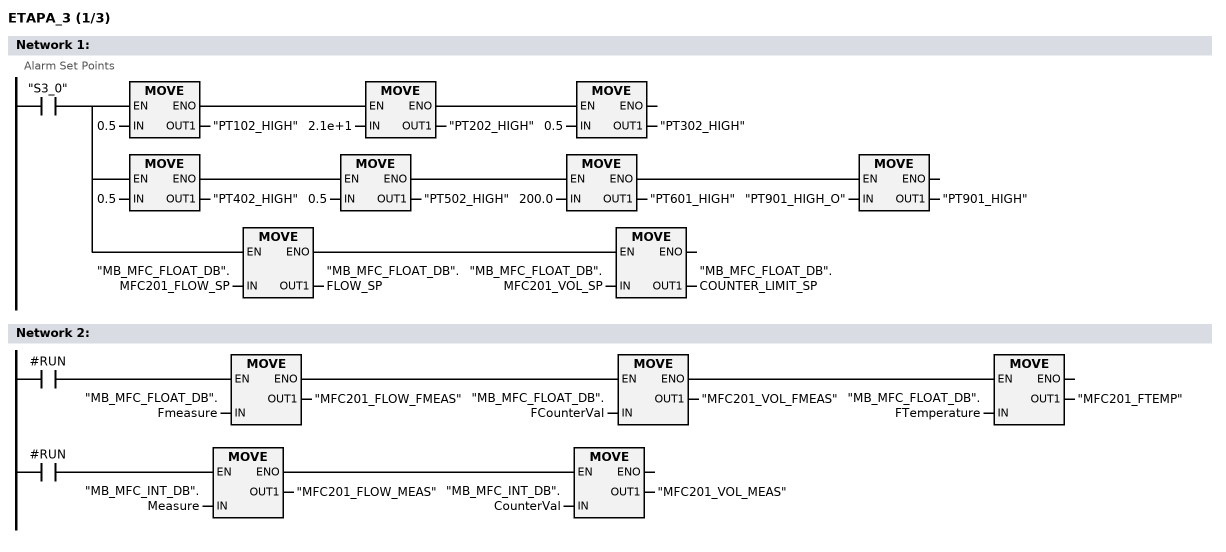
   RUNG wire#powerrail
      Contact( "S3_0" )
      wire#w1
      { S7_GenerateENO := "TRUE" } Move(in := 0.5, out1 => "PT102_HIGH")
      { S7_GenerateENO := "TRUE" } Move(in := 2.1e+1, out1 => "PT202_HIGH")
      { S7_GenerateENO := "TRUE" } Move(in := 0.5, out1 => "PT302_HIGH")
   END_RUNG
   RUNG wire#w1
      { S7_GenerateENO := "TRUE" } Move(in := 0.5, out1 => "PT402_HIGH")
      { S7_GenerateENO := "TRUE" } Move(in := 0.5, out1 => "PT502_HIGH")
      { S7_GenerateENO := "TRUE" } Move(in := 200.0, out1 => "PT601_HIGH")
      { S7_GenerateENO := "TRUE" } Move(in := "PT901_HIGH_O", out1 => "PT901_HIGH")
   END_RUNG
   RUNG wire#w1
      Move(in := "MB_MFC_FLOAT_DB".MFC201_FLOW_SP, out1 => "MB_MFC_FLOAT_DB".FLOW_SP)
      Move(in := "MB_MFC_FLOAT_DB".MFC201_VOL_SP, out1 => "MB_MFC_FLOAT_DB".COUNTER_LIMIT_SP)
   END_RUNG
   // the same network as SCL:
   // ENO of a box is taken as its EN; it also drops when the box reports an error
   IF "S3_0" THEN
       "PT102_HIGH" := 0.5;
       "PT202_HIGH" := 2.1e+1;
       "PT302_HIGH" := 0.5;
       "PT402_HIGH" := 0.5;
       "PT502_HIGH" := 0.5;
       "PT601_HIGH" := 200.0;
       "PT901_HIGH" := "PT901_HIGH_O";
       "MB_MFC_FLOAT_DB".FLOW_SP := "MB_MFC_FLOAT_DB".MFC201_FLOW_SP;
       "MB_MFC_FLOAT_DB".COUNTER_LIMIT_SP := "MB_MFC_FLOAT_DB".MFC201_VOL_SP;
   END_IF;
END_REGION

REGION Network 2
   RUNG wire#powerrail
      Contact( #RUN )
      { S7_GenerateENO := "TRUE" } Move(in := "MB_MFC_FLOAT_DB".Fmeasure, out1 => "MFC201_FLOW_FMEAS")
      { S7_GenerateENO := "TRUE" } Move(in := "MB_MFC_FLOAT_DB".FCounterVal, out1 => "MFC201_VOL_FMEAS")
      { S7_GenerateENO := "TRUE" } Move(in := "MB_MFC_FLOAT_DB".FTemperature, out1 => "MFC201_FTEMP")
   END_RUNG
   RUNG wire#powerrail
      Contact( #RUN )
      { S7_GenerateENO := "TRUE" } Move(in := "MB_MFC_INT_DB".Measure, out1 => "MFC201_FLOW_MEAS")
      { S7_GenerateENO := "TRUE" } Move(in := "MB_MFC_INT_DB".CounterVal, out1 => "MFC201_VOL_MEAS")
   END_RUNG
   // the same network as SCL:
   // ENO of a box is taken as its EN; it also drops when the box reports an error
   IF #RUN THEN
       "MFC201_FLOW_FMEAS" := "MB_MFC_FLOAT_DB".Fmeasure;
       "MFC201_VOL_FMEAS" := "MB_MFC_FLOAT_DB".FCounterVal;
       "MFC201_FTEMP" := "MB_MFC_FLOAT_DB".FTemperature;
       "MFC201_FLOW_MEAS" := "MB_MFC_INT_DB".Measure;
       "MFC201_VOL_MEAS" := "MB_MFC_INT_DB".CounterVal;
   END_IF;
END_REGION

REGION Network 3
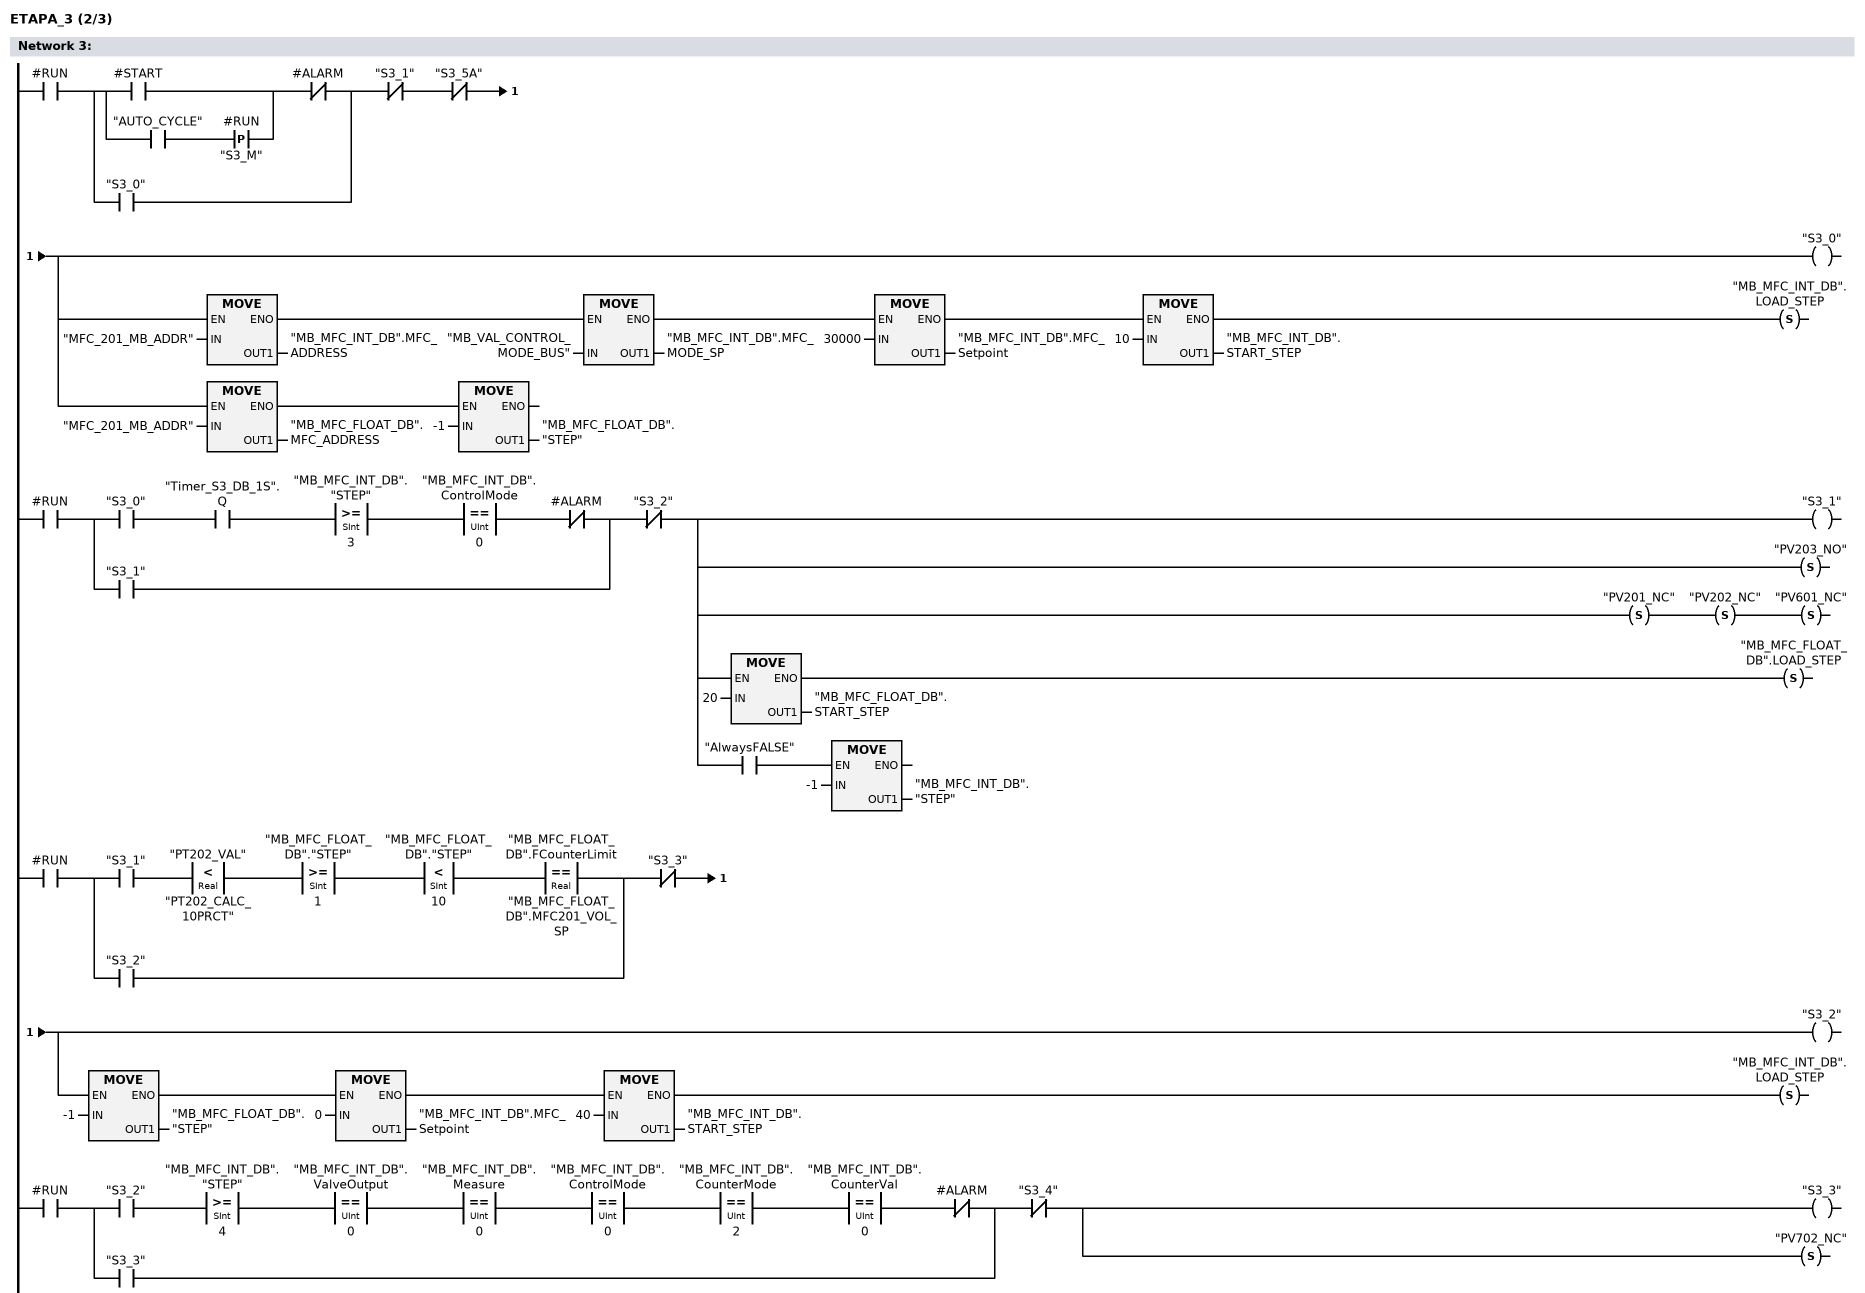
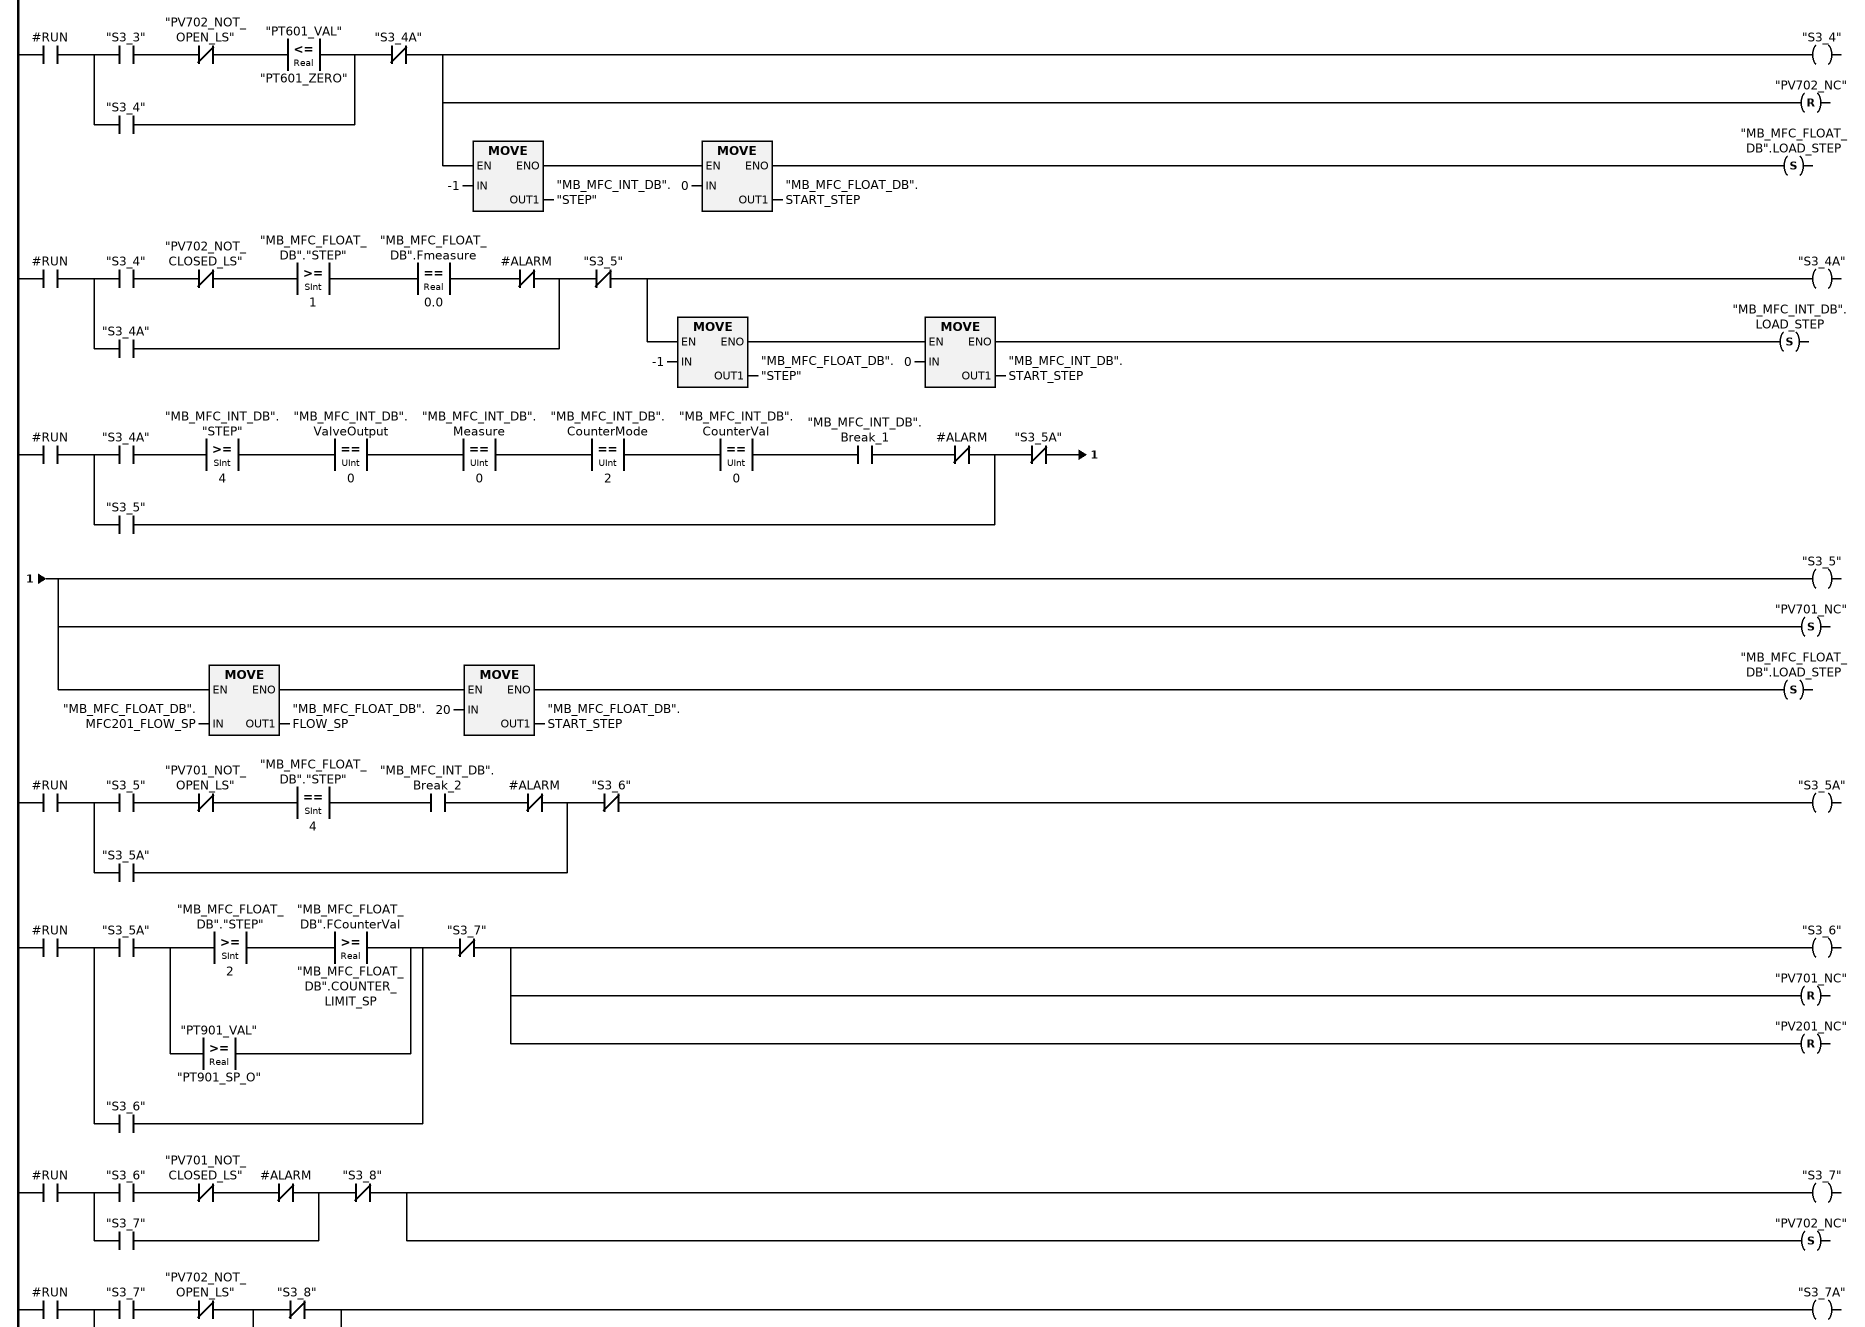
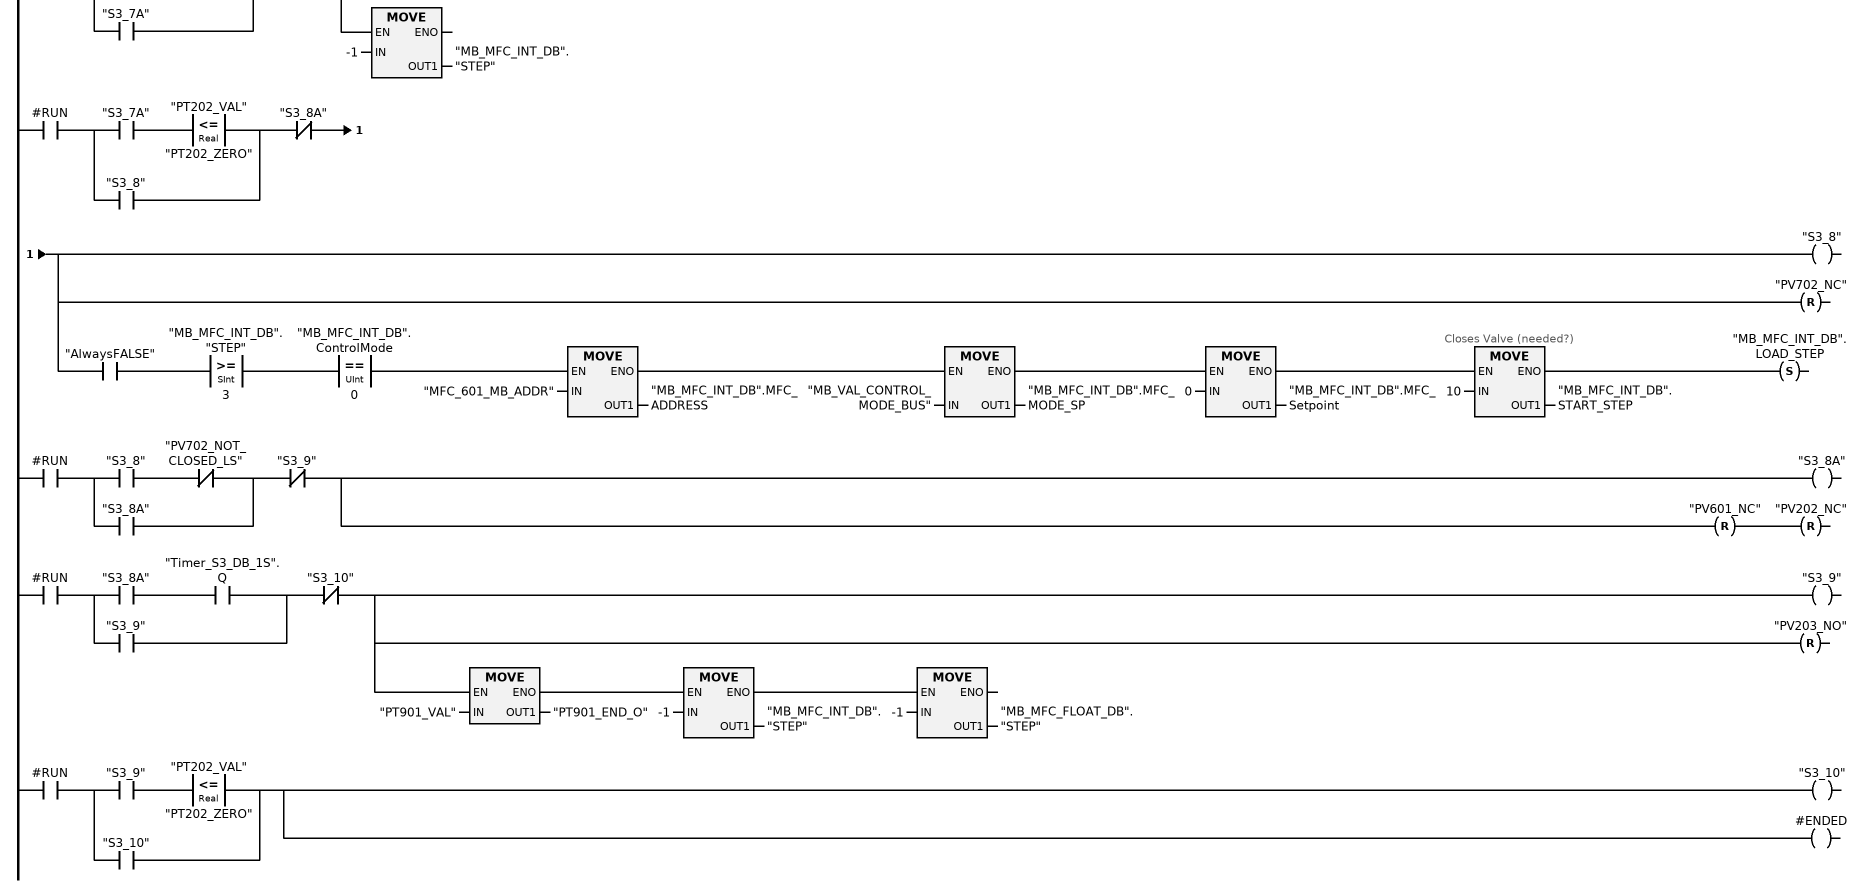
   RUNG wire#powerrail
      Contact( #RUN )
      wire#w1
      Contact( #START )
      wire#w2
      I_Contact( #ALARM )
      wire#w3
      I_Contact( "S3_1" )
      I_Contact( "S3_5A" )
      wire#w4
      Coil( "S3_0" )
   END_RUNG
   RUNG wire#w1
      Contact( "AUTO_CYCLE" )
      P_Contact(operand := #RUN, bit := "S3_M")
   END_RUNG wire#w2
   RUNG wire#w1
      Contact( "S3_0" )
   END_RUNG wire#w3
   RUNG wire#w4
      Move(in := "MFC_201_MB_ADDR", out1 => "MB_MFC_INT_DB".MFC_ADDRESS)
      Move(in := "MB_VAL_CONTROL_MODE_BUS", out1 => "MB_MFC_INT_DB".MFC_MODE_SP)
      Move(in := 30000, out1 => "MB_MFC_INT_DB".MFC_Setpoint)
      Move(in := 10, out1 => "MB_MFC_INT_DB".START_STEP)
      S_Coil( "MB_MFC_INT_DB".LOAD_STEP )
   END_RUNG
   RUNG wire#w4
      Move(in := "MFC_201_MB_ADDR", out1 => "MB_MFC_FLOAT_DB".MFC_ADDRESS)
      Move(in := -1, out1 => "MB_MFC_FLOAT_DB"."STEP")
   END_RUNG
   RUNG wire#powerrail
      Contact( #RUN )
      wire#w5
      Contact( "S3_0" )
      Contact( "Timer_S3_DB_1S".Q )
      { S7_Templates := "SrcType := SInt" } GE_Contact(in1 := "MB_MFC_INT_DB"."STEP", in2 := 3)
      { S7_Templates := "SrcType := UInt" } EQ_Contact(in1 := "MB_MFC_INT_DB".ControlMode, in2 := 0)
      I_Contact( #ALARM )
      wire#w6
      I_Contact( "S3_2" )
      wire#w7
      Coil( "S3_1" )
   END_RUNG
   RUNG wire#w5
      Contact( "S3_1" )
   END_RUNG wire#w6
   RUNG wire#w7
      S_Coil( "PV203_NO" )
   END_RUNG
   RUNG wire#w7
      S_Coil( "PV201_NC" )
      S_Coil( "PV202_NC" )
      S_Coil( "PV601_NC" )
   END_RUNG
   RUNG wire#w7
      Move(in := 20, out1 => "MB_MFC_FLOAT_DB".START_STEP)
      S_Coil( "MB_MFC_FLOAT_DB".LOAD_STEP )
   END_RUNG
   RUNG wire#w7
      Contact( "AlwaysFALSE" )
      Move(in := -1, out1 => "MB_MFC_INT_DB"."STEP")
   END_RUNG
   RUNG wire#powerrail
      Contact( #RUN )
      wire#w8
      Contact( "S3_1" )
      { S7_Templates := "SrcType := Real" } LT_Contact(in1 := "PT202_VAL", in2 := "PT202_CALC_10PRCT")
      { S7_Templates := "SrcType := SInt" } GE_Contact(in1 := "MB_MFC_FLOAT_DB"."STEP", in2 := 1)
      { S7_Templates := "SrcType := SInt" } LT_Contact(in1 := "MB_MFC_FLOAT_DB"."STEP", in2 := 10)
      { S7_Templates := "SrcType := Real" } EQ_Contact(in1 := "MB_MFC_FLOAT_DB".FCounterLimit, in2 := "MB_MFC_FLOAT_DB".MFC201_VOL_SP)
      wire#w9
      I_Contact( "S3_3" )
      wire#w10
      Coil( "S3_2" )
   END_RUNG
   RUNG wire#w8
      Contact( "S3_2" )
   END_RUNG wire#w9
   RUNG wire#w10
      Move(in := -1, out1 => "MB_MFC_FLOAT_DB"."STEP")
      Move(in := 0, out1 => "MB_MFC_INT_DB".MFC_Setpoint)
      Move(in := 40, out1 => "MB_MFC_INT_DB".START_STEP)
      S_Coil( "MB_MFC_INT_DB".LOAD_STEP )
   END_RUNG
   RUNG wire#powerrail
      Contact( #RUN )
      wire#w11
      Contact( "S3_2" )
      { S7_Templates := "SrcType := SInt" } GE_Contact(in1 := "MB_MFC_INT_DB"."STEP", in2 := 4)
      { S7_Templates := "SrcType := UInt" } EQ_Contact(in1 := "MB_MFC_INT_DB".ValveOutput, in2 := 0)
      { S7_Templates := "SrcType := UInt" } EQ_Contact(in1 := "MB_MFC_INT_DB".Measure, in2 := 0)
      { S7_Templates := "SrcType := UInt" } EQ_Contact(in1 := "MB_MFC_INT_DB".ControlMode, in2 := 0)
      { S7_Templates := "SrcType := UInt" } EQ_Contact(in1 := "MB_MFC_INT_DB".CounterMode, in2 := 2)
      { S7_Templates := "SrcType := UInt" } EQ_Contact(in1 := "MB_MFC_INT_DB".CounterVal, in2 := 0)
      I_Contact( #ALARM )
      wire#w12
      I_Contact( "S3_4" )
      wire#w13
      Coil( "S3_3" )
   END_RUNG
   RUNG wire#w11
      Contact( "S3_3" )
   END_RUNG wire#w12
   RUNG wire#w13
      S_Coil( "PV702_NC" )
   END_RUNG
   RUNG wire#powerrail
      Contact( #RUN )
      wire#w14
      Contact( "S3_3" )
      I_Contact( "PV702_NOT_OPEN_LS" )
      { S7_Templates := "SrcType := Real" } LE_Contact(in1 := "PT601_VAL", in2 := "PT601_ZERO")
      wire#w15
      I_Contact( "S3_4A" )
      wire#w16
      Coil( "S3_4" )
   END_RUNG
   RUNG wire#w14
      Contact( "S3_4" )
   END_RUNG wire#w15
   RUNG wire#w16
      R_Coil( "PV702_NC" )
   END_RUNG
   RUNG wire#w16
      Move(in := -1, out1 => "MB_MFC_INT_DB"."STEP")
      Move(in := 0, out1 => "MB_MFC_FLOAT_DB".START_STEP)
      S_Coil( "MB_MFC_FLOAT_DB".LOAD_STEP )
   END_RUNG
   RUNG wire#powerrail
      Contact( #RUN )
      wire#w17
      Contact( "S3_4" )
      I_Contact( "PV702_NOT_CLOSED_LS" )
      { S7_Templates := "SrcType := SInt" } GE_Contact(in1 := "MB_MFC_FLOAT_DB"."STEP", in2 := 1)
      { S7_Templates := "SrcType := Real" } EQ_Contact(in1 := "MB_MFC_FLOAT_DB".Fmeasure, in2 := 0.0)
      I_Contact( #ALARM )
      wire#w18
      I_Contact( "S3_5" )
      wire#w19
      Coil( "S3_4A" )
   END_RUNG
   RUNG wire#w17
      Contact( "S3_4A" )
   END_RUNG wire#w18
   RUNG wire#w19
      Move(in := -1, out1 => "MB_MFC_FLOAT_DB"."STEP")
      Move(in := 0, out1 => "MB_MFC_INT_DB".START_STEP)
      S_Coil( "MB_MFC_INT_DB".LOAD_STEP )
   END_RUNG
   RUNG wire#powerrail
      Contact( #RUN )
      wire#w20
      Contact( "S3_4A" )
      { S7_Templates := "SrcType := SInt" } GE_Contact(in1 := "MB_MFC_INT_DB"."STEP", in2 := 4)
      { S7_Templates := "SrcType := UInt" } EQ_Contact(in1 := "MB_MFC_INT_DB".ValveOutput, in2 := 0)
      { S7_Templates := "SrcType := UInt" } EQ_Contact(in1 := "MB_MFC_INT_DB".Measure, in2 := 0)
      { S7_Templates := "SrcType := UInt" } EQ_Contact(in1 := "MB_MFC_INT_DB".CounterMode, in2 := 2)
      { S7_Templates := "SrcType := UInt" } EQ_Contact(in1 := "MB_MFC_INT_DB".CounterVal, in2 := 0)
      Contact( "MB_MFC_INT_DB".Break_1 )
      I_Contact( #ALARM )
      wire#w21
      I_Contact( "S3_5A" )
      wire#w22
      Coil( "S3_5" )
   END_RUNG
   RUNG wire#w20
      Contact( "S3_5" )
   END_RUNG wire#w21
   RUNG wire#w22
      S_Coil( "PV701_NC" )
   END_RUNG
   RUNG wire#w22
      Move(in := "MB_MFC_FLOAT_DB".MFC201_FLOW_SP, out1 => "MB_MFC_FLOAT_DB".FLOW_SP)
      Move(in := 20, out1 => "MB_MFC_FLOAT_DB".START_STEP)
      S_Coil( "MB_MFC_FLOAT_DB".LOAD_STEP )
   END_RUNG
   RUNG wire#powerrail
      Contact( #RUN )
      wire#w23
      Contact( "S3_5" )
      I_Contact( "PV701_NOT_OPEN_LS" )
      { S7_Templates := "SrcType := SInt" } EQ_Contact(in1 := "MB_MFC_FLOAT_DB"."STEP", in2 := 4)
      Contact( "MB_MFC_INT_DB".Break_2 )
      I_Contact( #ALARM )
      wire#w24
      I_Contact( "S3_6" )
      Coil( "S3_5A" )
   END_RUNG
   RUNG wire#w23
      Contact( "S3_5A" )
   END_RUNG wire#w24
   RUNG wire#powerrail
      Contact( #RUN )
      wire#w25
      Contact( "S3_5A" )
      wire#w26
      { S7_Templates := "SrcType := SInt" } GE_Contact(in1 := "MB_MFC_FLOAT_DB"."STEP", in2 := 2)
      { S7_Templates := "SrcType := Real" } GE_Contact(in1 := "MB_MFC_FLOAT_DB".FCounterVal, in2 := "MB_MFC_FLOAT_DB".COUNTER_LIMIT_SP)
      wire#w27
      I_Contact( "S3_7" )
      wire#w28
      Coil( "S3_6" )
   END_RUNG
   RUNG wire#w26
      { S7_Templates := "SrcType := Real" } GE_Contact(in1 := "PT901_VAL", in2 := "PT901_SP_O")
   END_RUNG wire#w27
   RUNG wire#w25
      Contact( "S3_6" )
   END_RUNG wire#w27
   RUNG wire#w28
      R_Coil( "PV701_NC" )
   END_RUNG
   RUNG wire#w28
      R_Coil( "PV201_NC" )
   END_RUNG
   RUNG wire#powerrail
      Contact( #RUN )
      wire#w29
      Contact( "S3_6" )
      I_Contact( "PV701_NOT_CLOSED_LS" )
      I_Contact( #ALARM )
      wire#w30
      I_Contact( "S3_8" )
      wire#w31
      Coil( "S3_7" )
   END_RUNG
   RUNG wire#w29
      Contact( "S3_7" )
   END_RUNG wire#w30
   RUNG wire#w31
      S_Coil( "PV702_NC" )
   END_RUNG
   RUNG wire#powerrail
      Contact( #RUN )
      wire#w32
      Contact( "S3_7" )
      I_Contact( "PV702_NOT_OPEN_LS" )
      wire#w33
      I_Contact( "S3_8" )
      wire#w34
      Coil( "S3_7A" )
   END_RUNG
   RUNG wire#w32
      Contact( "S3_7A" )
   END_RUNG wire#w33
   RUNG wire#w34
      Move(in := -1, out1 => "MB_MFC_INT_DB"."STEP")
   END_RUNG
   RUNG wire#powerrail
      Contact( #RUN )
      wire#w35
      Contact( "S3_7A" )
      { S7_Templates := "SrcType := Real" } LE_Contact(in1 := "PT202_VAL", in2 := "PT202_ZERO")
      wire#w36
      I_Contact( "S3_8A" )
      wire#w37
      Coil( "S3_8" )
   END_RUNG
   RUNG wire#w35
      Contact( "S3_8" )
   END_RUNG wire#w36
   RUNG wire#w37
      R_Coil( "PV702_NC" )
   END_RUNG
   RUNG wire#w37
      Contact( "AlwaysFALSE" )
      { S7_Templates := "SrcType := SInt" } GE_Contact(in1 := "MB_MFC_INT_DB"."STEP", in2 := 3)
      { S7_Templates := "SrcType := UInt" } EQ_Contact(in1 := "MB_MFC_INT_DB".ControlMode, in2 := 0)
      Move(in := "MFC_601_MB_ADDR", out1 => "MB_MFC_INT_DB".MFC_ADDRESS)
      Move(in := "MB_VAL_CONTROL_MODE_BUS", out1 => "MB_MFC_INT_DB".MFC_MODE_SP)
      Move(in := 0, out1 => "MB_MFC_INT_DB".MFC_Setpoint)
      Move(in := 10, out1 => "MB_MFC_INT_DB".START_STEP)   // Closes Valve (needed?)
      S_Coil( "MB_MFC_INT_DB".LOAD_STEP )
   END_RUNG
   RUNG wire#powerrail
      Contact( #RUN )
      wire#w38
      Contact( "S3_8" )
      I_Contact( "PV702_NOT_CLOSED_LS" )
      wire#w39
      I_Contact( "S3_9" )
      wire#w40
      Coil( "S3_8A" )
   END_RUNG
   RUNG wire#w38
      Contact( "S3_8A" )
   END_RUNG wire#w39
   RUNG wire#w40
      R_Coil( "PV601_NC" )
      R_Coil( "PV202_NC" )
   END_RUNG
   RUNG wire#powerrail
      Contact( #RUN )
      wire#w41
      Contact( "S3_8A" )
      Contact( "Timer_S3_DB_1S".Q )
      wire#w42
      I_Contact( "S3_10" )
      wire#w43
      Coil( "S3_9" )
   END_RUNG
   RUNG wire#w41
      Contact( "S3_9" )
   END_RUNG wire#w42
   RUNG wire#w43
      R_Coil( "PV203_NO" )
   END_RUNG
   RUNG wire#w43
      { S7_GenerateENO := "TRUE" } Move(in := "PT901_VAL", out1 => "PT901_END_O")
      Move(in := -1, out1 => "MB_MFC_INT_DB"."STEP")
      Move(in := -1, out1 => "MB_MFC_FLOAT_DB"."STEP")
   END_RUNG
   RUNG wire#powerrail
      Contact( #RUN )
      wire#w44
      Contact( "S3_9" )
      { S7_Templates := "SrcType := Real" } LE_Contact(in1 := "PT202_VAL", in2 := "PT202_ZERO")
      wire#w45
      Coil( "S3_10" )
   END_RUNG
   RUNG wire#w44
      Contact( "S3_10" )
   END_RUNG wire#w45
   RUNG wire#w45
      Coil( #ENDED )
   END_RUNG
   // the same network as SCL:
   // ENO of a box is taken as its EN; it also drops when the box reports an error
   #_w1 := #RUN AND "AUTO_CYCLE" AND #RUN AND NOT "S3_M";   // rising edge of #RUN
   "S3_M" := #RUN;
   "S3_0" := ((((#RUN AND #START) OR #_w1) AND NOT #ALARM) OR (#RUN AND "S3_0")) AND NOT "S3_1" AND NOT "S3_5A";
   IF "S3_0" THEN
       "MB_MFC_INT_DB".MFC_ADDRESS := "MFC_201_MB_ADDR";
       "MB_MFC_INT_DB".MFC_MODE_SP := "MB_VAL_CONTROL_MODE_BUS";
       "MB_MFC_INT_DB".MFC_Setpoint := 30000;
       "MB_MFC_INT_DB".START_STEP := 10;
       "MB_MFC_INT_DB".LOAD_STEP := TRUE;
       "MB_MFC_FLOAT_DB".MFC_ADDRESS := "MFC_201_MB_ADDR";
       "MB_MFC_FLOAT_DB"."STEP" := -1;
   END_IF;
   "S3_1" := #RUN AND (("S3_0" AND "Timer_S3_DB_1S".Q AND ("MB_MFC_INT_DB"."STEP" >= 3) AND ("MB_MFC_INT_DB".ControlMode = 0) AND NOT #ALARM) OR "S3_1") AND NOT "S3_2";
   IF "S3_1" THEN
       "PV203_NO" := TRUE;
       "PV201_NC" := TRUE;
       "PV202_NC" := TRUE;
       "PV601_NC" := TRUE;
       "MB_MFC_FLOAT_DB".START_STEP := 20;
       "MB_MFC_FLOAT_DB".LOAD_STEP := TRUE;
   END_IF;
   IF "S3_1" AND "AlwaysFALSE" THEN "MB_MFC_INT_DB"."STEP" := -1; END_IF;
   "S3_2" := #RUN AND (("S3_1" AND ("PT202_VAL" < "PT202_CALC_10PRCT") AND ("MB_MFC_FLOAT_DB"."STEP" >= 1) AND ("MB_MFC_FLOAT_DB"."STEP" < 10) AND ("MB_MFC_FLOAT_DB".FCounterLimit = "MB_MFC_FLOAT_DB".MFC201_VOL_SP)) OR "S3_2") AND NOT "S3_3";
   IF "S3_2" THEN
       "MB_MFC_FLOAT_DB"."STEP" := -1;
       "MB_MFC_INT_DB".MFC_Setpoint := 0;
       "MB_MFC_INT_DB".START_STEP := 40;
       "MB_MFC_INT_DB".LOAD_STEP := TRUE;
   END_IF;
   "S3_3" := #RUN AND (("S3_2" AND ("MB_MFC_INT_DB"."STEP" >= 4) AND ("MB_MFC_INT_DB".ValveOutput = 0) AND ("MB_MFC_INT_DB".Measure = 0) AND ("MB_MFC_INT_DB".ControlMode = 0) AND ("MB_MFC_INT_DB".CounterMode = 2) AND ("MB_MFC_INT_DB".CounterVal = 0) AND NOT #ALARM) OR "S3_3") AND NOT "S3_4";
   IF "S3_3" THEN "PV702_NC" := TRUE; END_IF;
   "S3_4" := #RUN AND (("S3_3" AND NOT "PV702_NOT_OPEN_LS" AND ("PT601_VAL" <= "PT601_ZERO")) OR "S3_4") AND NOT "S3_4A";
   IF "S3_4" THEN
       "PV702_NC" := FALSE;
       "MB_MFC_INT_DB"."STEP" := -1;
       "MB_MFC_FLOAT_DB".START_STEP := 0;
       "MB_MFC_FLOAT_DB".LOAD_STEP := TRUE;
   END_IF;
   "S3_4A" := #RUN AND (("S3_4" AND NOT "PV702_NOT_CLOSED_LS" AND ("MB_MFC_FLOAT_DB"."STEP" >= 1) AND ("MB_MFC_FLOAT_DB".Fmeasure = 0.0) AND NOT #ALARM) OR "S3_4A") AND NOT "S3_5";
   IF "S3_4A" THEN
       "MB_MFC_FLOAT_DB"."STEP" := -1;
       "MB_MFC_INT_DB".START_STEP := 0;
       "MB_MFC_INT_DB".LOAD_STEP := TRUE;
   END_IF;
   "S3_5" := #RUN AND (("S3_4A" AND ("MB_MFC_INT_DB"."STEP" >= 4) AND ("MB_MFC_INT_DB".ValveOutput = 0) AND ("MB_MFC_INT_DB".Measure = 0) AND ("MB_MFC_INT_DB".CounterMode = 2) AND ("MB_MFC_INT_DB".CounterVal = 0) AND "MB_MFC_INT_DB".Break_1 AND NOT #ALARM) OR "S3_5") AND NOT "S3_5A";
   IF "S3_5" THEN
       "PV701_NC" := TRUE;
       "MB_MFC_FLOAT_DB".FLOW_SP := "MB_MFC_FLOAT_DB".MFC201_FLOW_SP;
       "MB_MFC_FLOAT_DB".START_STEP := 20;
       "MB_MFC_FLOAT_DB".LOAD_STEP := TRUE;
   END_IF;
   "S3_5A" := #RUN AND (("S3_5" AND NOT "PV701_NOT_OPEN_LS" AND ("MB_MFC_FLOAT_DB"."STEP" = 4) AND "MB_MFC_INT_DB".Break_2 AND NOT #ALARM) OR "S3_5A") AND NOT "S3_6";
   "S3_6" := #RUN AND (("S3_5A" AND ((("MB_MFC_FLOAT_DB"."STEP" >= 2) AND ("MB_MFC_FLOAT_DB".FCounterVal >= "MB_MFC_FLOAT_DB".COUNTER_LIMIT_SP)) OR ("PT901_VAL" >= "PT901_SP_O"))) OR "S3_6") AND NOT "S3_7";
   IF "S3_6" THEN
       "PV701_NC" := FALSE;
       "PV201_NC" := FALSE;
   END_IF;
   "S3_7" := #RUN AND (("S3_6" AND NOT "PV701_NOT_CLOSED_LS" AND NOT #ALARM) OR "S3_7") AND NOT "S3_8";
   IF "S3_7" THEN "PV702_NC" := TRUE; END_IF;
   "S3_7A" := #RUN AND (("S3_7" AND NOT "PV702_NOT_OPEN_LS") OR "S3_7A") AND NOT "S3_8";
   IF "S3_7A" THEN "MB_MFC_INT_DB"."STEP" := -1; END_IF;
   "S3_8" := #RUN AND (("S3_7A" AND ("PT202_VAL" <= "PT202_ZERO")) OR "S3_8") AND NOT "S3_8A";
   IF "S3_8" THEN "PV702_NC" := FALSE; END_IF;
   IF "S3_8" AND "AlwaysFALSE" AND ("MB_MFC_INT_DB"."STEP" >= 3) AND ("MB_MFC_INT_DB".ControlMode = 0) THEN
       "MB_MFC_INT_DB".MFC_ADDRESS := "MFC_601_MB_ADDR";
       "MB_MFC_INT_DB".MFC_MODE_SP := "MB_VAL_CONTROL_MODE_BUS";
       "MB_MFC_INT_DB".MFC_Setpoint := 0;
       "MB_MFC_INT_DB".START_STEP := 10;   // Closes Valve (needed?)
       "MB_MFC_INT_DB".LOAD_STEP := TRUE;
   END_IF;
   "S3_8A" := #RUN AND (("S3_8" AND NOT "PV702_NOT_CLOSED_LS") OR "S3_8A") AND NOT "S3_9";
   IF "S3_8A" THEN
       "PV601_NC" := FALSE;
       "PV202_NC" := FALSE;
   END_IF;
   "S3_9" := #RUN AND (("S3_8A" AND "Timer_S3_DB_1S".Q) OR "S3_9") AND NOT "S3_10";
   IF "S3_9" THEN
       "PV203_NO" := FALSE;
       "PT901_END_O" := "PT901_VAL";
       "MB_MFC_INT_DB"."STEP" := -1;
       "MB_MFC_FLOAT_DB"."STEP" := -1;
   END_IF;
   "S3_10" := #RUN AND (("S3_9" AND ("PT202_VAL" <= "PT202_ZERO")) OR "S3_10");
   #ENDED := "S3_10";
END_REGION

REGION Network 4
   // Timers
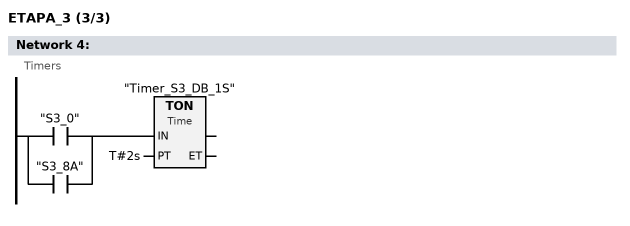
   "Timer_S3_DB_1S".TON(IN := "S3_0" OR "S3_8A", PT := T#2s);
END_REGION
END_FUNCTION

FUNCTION "ETAPA_4" : Void   // FC5, LAD
{ S7_Optimized_Access := 'FALSE' }
VERSION : 0.1
// Injecao de Helio 1, Controlo por Volume
   VAR_TEMP   // added for the SCL form of the ladder/FBD networks
      _w1 : Bool;
   END_VAR
BEGIN

REGION Network 1
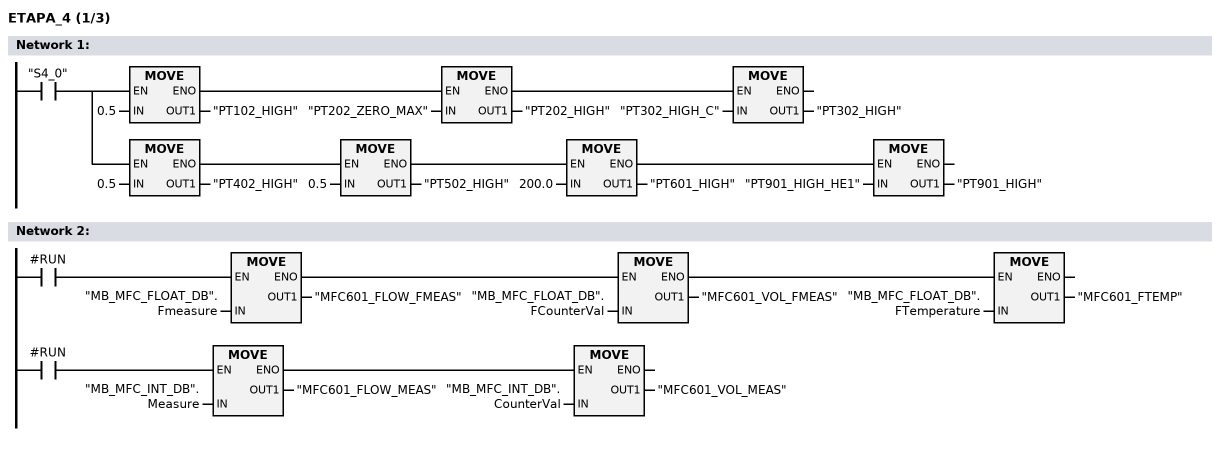
   RUNG wire#powerrail
      Contact( "S4_0" )
      wire#w1
      { S7_GenerateENO := "TRUE" } Move(in := 0.5, out1 => "PT102_HIGH")
      { S7_GenerateENO := "TRUE" } Move(in := "PT202_ZERO_MAX", out1 => "PT202_HIGH")
      { S7_GenerateENO := "TRUE" } Move(in := "PT302_HIGH_C", out1 => "PT302_HIGH")
   END_RUNG
   RUNG wire#w1
      { S7_GenerateENO := "TRUE" } Move(in := 0.5, out1 => "PT402_HIGH")
      { S7_GenerateENO := "TRUE" } Move(in := 0.5, out1 => "PT502_HIGH")
      { S7_GenerateENO := "TRUE" } Move(in := 200.0, out1 => "PT601_HIGH")
      { S7_GenerateENO := "TRUE" } Move(in := "PT901_HIGH_HE1", out1 => "PT901_HIGH")
   END_RUNG
   // the same network as SCL:
   // ENO of a box is taken as its EN; it also drops when the box reports an error
   IF "S4_0" THEN
       "PT102_HIGH" := 0.5;
       "PT202_HIGH" := "PT202_ZERO_MAX";
       "PT302_HIGH" := "PT302_HIGH_C";
       "PT402_HIGH" := 0.5;
       "PT502_HIGH" := 0.5;
       "PT601_HIGH" := 200.0;
       "PT901_HIGH" := "PT901_HIGH_HE1";
   END_IF;
END_REGION

REGION Network 2
   RUNG wire#powerrail
      Contact( #RUN )
      { S7_GenerateENO := "TRUE" } Move(in := "MB_MFC_FLOAT_DB".Fmeasure, out1 => "MFC601_FLOW_FMEAS")
      { S7_GenerateENO := "TRUE" } Move(in := "MB_MFC_FLOAT_DB".FCounterVal, out1 => "MFC601_VOL_FMEAS")
      { S7_GenerateENO := "TRUE" } Move(in := "MB_MFC_FLOAT_DB".FTemperature, out1 => "MFC601_FTEMP")
   END_RUNG
   RUNG wire#powerrail
      Contact( #RUN )
      { S7_GenerateENO := "TRUE" } Move(in := "MB_MFC_INT_DB".Measure, out1 => "MFC601_FLOW_MEAS")
      { S7_GenerateENO := "TRUE" } Move(in := "MB_MFC_INT_DB".CounterVal, out1 => "MFC601_VOL_MEAS")
   END_RUNG
   // the same network as SCL:
   // ENO of a box is taken as its EN; it also drops when the box reports an error
   IF #RUN THEN
       "MFC601_FLOW_FMEAS" := "MB_MFC_FLOAT_DB".Fmeasure;
       "MFC601_VOL_FMEAS" := "MB_MFC_FLOAT_DB".FCounterVal;
       "MFC601_FTEMP" := "MB_MFC_FLOAT_DB".FTemperature;
       "MFC601_FLOW_MEAS" := "MB_MFC_INT_DB".Measure;
       "MFC601_VOL_MEAS" := "MB_MFC_INT_DB".CounterVal;
   END_IF;
END_REGION

REGION Network 3